TYPE "UDT_SDC_EMS_TS_COM"
VERSION : 0.1
   STRUCT
      VAL : "UDT_SDC_TS_IF_COMMAND_VAL";
      BIT : "UDT_SDC_TS_IF_COMMAND_BIT";
      FKT_SET : "UDT_SDC_EMS_FKT_BITs";
      FKT_RESET : "UDT_SDC_EMS_FKT_BITs";
   END_STRUCT;
END_TYPE

TYPE "UDT_EMS_IF_Q_STAT"
VERSION : 0.1
   STRUCT
      LIFE_BIT : Bool;   // Lebensbit / Heartbeat
      ER_SUM : Bool;   // Sammelfehler / Summaryerror
      IR_MAN : Bool;   // EMS in Handbetrieb / EMS in manual mode (IR)
      ER_RESET : Bool;   // Störung quittieren / Error reset (IR)
      HOIST_CLEAR : Bool;   // Hub über/in Sollpos und Bereit ohne Störung / Hoist above position and no error
      POS_START_X : Bool;   // Fahrantrieb positioniert / Drive positioning started
      ALWAYS_ONE : Bool;   // immer "1" / Always "1"
      H_DISABLED : Bool;   // Hub gesperrt / Hoist disabled
      D_FWD : Bool;   // Fahrantrieb fährt vorwärts / Drive moves forwards
      D_RWD : Bool;   // Fahrantrieb fährt rückwärts / Drive moves reward
      bit12 : Bool;   // Reserve / spare
      D_IN_POS : Bool;   // Fahrantrieb in Position / Drive in Position
      H_UP : Bool;   // Hub hebt / Hoist raises
      H_DOWN : Bool;   // Hub senkt / Hoist lowers
      H_IN_POS : Bool;   // Hub in Position / Hoist in position
      H_IN_TOPPOS : Bool;   // Hub in oberster Position / Hoist in top position
      bit2_0 : Bool;   // Schwenkantrieb fährt + / Tilt moves clockwise
      bit2_1 : Bool;   // Schwenkantrieb fährt - / Tilt moves counterclockwise
      bit2_2 : Bool;   // Hub in oberster Position / Tilt in position
      bit2_3 : Bool;   // Hub in Grundstellung / Tilt in home position
      IN_BOTPOS : Bool;   // Hub in unterster Position / Hoist In bottom Position (min) (with Tiltposition)
      bit2_5 : Bool;   // Reserve / spare
      bit2_6 : Bool;   // Reserve / spare
      bit2_7 : Bool;   // Reserve / spare
      MESS_ACT : Bool;   // Störnummer ist eine Meldung / Error No is a Message
      MESS_POS : Bool;   // Reserve / spare
      bit3_2 : Bool;   // Reserve / spare
      bit3_3 : Bool;   // Reserve / spare
      bit3_4 : Bool;   // Reserve / spare
      bit3_5 : Bool;   // Reserve / spare
      bit3_6 : Bool;   // Reserve / spare
      DATA_TRANS : Bool;   // Datentransfer ist aktiv / Data Transfer aktiv
   END_STRUCT;
END_TYPE

TYPE "UDT_EMS_IF_I_CONTR"
VERSION : 0.1
   STRUCT
      LIFE_BIT : Bool;   // Lebensbit / Heartbeat
      ER_SDC : Bool;   // Sammelfehler / Summaryerror
      H_EMERG : Bool;   // Hubantrieb Notbetrieb / Hoist Emergency mode
      Spare_0_3 : Bool;   // Schwenkantrieb Notbetrieb / Tilt Emergency mode
      LAMP_TEST : Bool;   // Lampentest / Lamp Test
      VAC_CLEAN : Bool;   // EMS mit Staubsauger / EMS with vac cleaner
      SYNCH : Bool;   // Synchronbetrieb / Control distance, synchronous area
      DATA_TRANS : Bool;   // Datentransfer ist aktiv / Data Transfer aktiv
      ER_RESET : Bool;   // Störung quittieren / Error reset
      AUTO : Bool;   // 1 = Automatikbetrieb / Automatic mode in section
      MAN : Bool;   // 1 = Handbetrieb / Manual mode in section
      D_C_BREAK : Bool;   // Fahrantrieb Befehl Bremse lüften / DRIVE Command release Break
      H_C_BREAK : Bool;   // Hubantrieb Befehl Bremse lüften / HOIST Command release Break
      D_EMERG_FC : Bool;   // Fahrantrieb Notbetrieb 1 Motor / DRIVE Emergency mode Frequencyconverter 1 Motor
      INC_TOL_POS : Bool;   // Schwenkantrieb Notbetrieb 1 Motor / TILT Emergency mode Frequencyconverter 1 Motor
      E_STOP : Bool;   // "1"Not-Halt / Emergency stop from Interface
      D_C_FWD : Bool;   // Fahrantrieb Befehl vorwärts / DRIVE Command forward
      D_C_RWD : Bool;   // Fahrantrieb Befehl rückwärts / DRIVE Command reward
      D_C_BSP : Bool;   // Fahrantrieb Befehl weiter fahren / DRIVE Command bridge stop position
      Spare_2_3 : Bool;   // Reserve / spare
      IR_noEMSnumber : Bool;   // Schwenkantrieb Befehl + / TILT Command clockwise
      IR_noLogin : Bool;   // Schwenkantrieb Befehl - / TILT Command counterclockwise
      BYP_scalance_PN_error : Bool;   // Schwenkantrieb Befehl positionieren / TILT Command positioning
      Spare_2_7 : Bool;   // Schwenkantrieb Befehl fahren in Grundstellung / TILT Command to home position, high priority
      H_C_UP : Bool;   // Hubantrieb Befehl heben / HOIST Command raise without positioning
      H_C_DOWN : Bool;   // Hubantrieb Befehl senken / HOIST Command lower without positioning
      H_C_POS : Bool;   // Hubantrieb Befehl positionieren / HOIST Command hoist positioning
      H_C_TOP : Bool;   // Hubantrieb Befehl fahren in oberste Position / HOIST Command Raise to top position, high priority
      H_EN : Bool;   // Hub-Schwenkfreigabe / HOIST-TILT enable
      H_BYP_ROPE : Bool;   // Überbrücken Seilkontrolle / Bypass monitoring of rope
      Spare_3_6 : Bool;   // Reserve / spare
      H_BYP_REF_INI : Bool;   // Überbrücken Kontrolle Referenzinitiator (nicht safety) / No monitoring of reference initiator (non safety)
   END_STRUCT;
END_TYPE

TYPE "UDT_SDC_TS_IF_COMMAND_BIT"
AUTHOR : SIEMENS
FAMILY : FT
NAME : SDC_BIT
VERSION : 2.0
   STRUCT
      ER_RESET : Bool;   // Error Reset
      AUTO : Bool;   // 1 = Automatik in Sektion
      MAN : Bool;   // 1 = Handbetrieb in Sektion
      Spare_0_3 : Bool;   // Reserve
      Spare_0_4 : Bool;   // Reserve
      E_STOP : Bool;   // "1" -> NotAus von Interface (system PLC)
      Spare_0_6 : Bool;   // Reserve
      Spare_0_7 : Bool;   // Reserve
      D_C_FWD : Bool;   // Fahrantrieb Kommando vorwärts
      D_C_RWD : Bool;   // Fahrantrieb Kommando rückwärts
      D_C_BSP : Bool;   // Fahrantrieb Kommando Überbrückung Stopp-Position
      D_C_V1 : Bool;   // Fahrantrieb Kommando Geschwindigkeit 1
      D_C_V2 : Bool;   // Fahrantrieb Kommando Geschwindigkeit 2
      D_C_V_VAR : Bool;   // Fahrantrieb Kommando variabler Geschwindigkeit
      D_C_BEFOR_POS : Bool;   // Fahrantrieb Kommando Freigabe vor Stop-Position
      D_C_AFTER_POS : Bool;   // Fahrantrieb Kommando Freigabe nach Stop-Position
      H_C_RAISE : Bool;   // Hubantrieb Kommando aufwärts
      H_C_LOWER : Bool;   // Hubantrieb Kommando abwärts
      H_C_POS : Bool;   // Hubantrieb Kommando Positionieren
      H_C_POS1 : Bool;   // Hubantrieb Kommando Offset 1
      H_C_POS2 : Bool;   // Hubantrieb Kommando Offset 2
      H_C_POS3 : Bool;   // Hubantrieb Kommando Offset 3
      H_C_POS4 : Bool;   // Hubantrieb Kommando Offset 4
      H_C_TOP : Bool;   // Hubantrieb Kommando nach Top Position, hohe Priorität
      H_BYP_ROPE : Bool;   // Hubantrieb Überbrücken Seilkontrolle
      Spare_3_1 : Bool;   // Reserve
      H_BYP_REF_INI : Bool;   // Hubantrieb Überbrücken Kontrolle Referenzinitiator (nicht safety)
      H_C_SLOW : Bool;   // Hubantrieb Kommando globaler Parameter langsam
      D_BYP_DIST_CONTR : Bool;   // Fahrantrieb Überbrücke Distanzkontrolle
      Spare_3_5 : Bool;   // Reserve
      Spare_3_6 : Bool;   // Reserve
      SET_PROF : Bool;   // setze Profile
   END_STRUCT;
END_TYPE

TYPE "UDT_SDC_TS_IF_COMMAND_VAL"
AUTHOR : SIEMENS
FAMILY : FT
NAME : SDC_VAL
VERSION : 1.6
   STRUCT
      PROFIL : Int;   // Profile
      D_SETSPEED : DInt;   // set value: drive speed (mm/min)
      D_POS_OFFS : Int;   // Antriebsposition offset
      H_POS_OFFS : Int;
   END_STRUCT;
END_TYPE

TYPE "UDT_SDC_TS_IF_STATUS_BIT"
AUTHOR : SIEMENS
FAMILY : FT
NAME : SDC_BIT
VERSION : 1.6
   STRUCT
      PRESENT : Bool;   // EMS vorhanden
      ERROR : Bool;   // Sammelstörung
      MAN_IR : Bool;   // EMS in Handbetrieb (Fernsteuerung)
      MORE_EMS_PRESENT : Bool;   // Mehr als 1 EMS in Sektion vorhanden
      ER_COMMAND : Bool;   // Fehlerhafte Befehle von System PLC
      W_DIST : Bool;   // Warnung Distanckontrolle ist aktiv
      Spare_0_6 : Bool;   // Warnung Auffahrsensor ist aktiv Reserve
      MESS_ACT : Bool;   // Störnummer ist eine Meldung / Error No is a Message
      D_MOVING : Bool;   // Fahrantrieb ist ein
      D_NOT_MOVING : Bool;   // Fahrantrieb ist aus
      H_MOVING : Bool;   // Hubantrieb ist ein
      H_NOT_MOVING : Bool;   // Hubantrieb ist aus
      X_MOVING : Bool;   // Reserve Antrieb ein
      X_NOT_MOVING : Bool;   // Reserve Antrieb aus
      D_IN_POS : Bool;   // Fahrantrieb in Position
      Spare_2_1 : Bool;   // Reserve
      D_BEFOR_POS : Bool;   // Fahrantrieb vor Stopposition
      D_AFTER_POS : Bool;   // Fahrantrieb nach Stopposition
      D_GR_AP1 : Bool;   // Fahrantrieb Barcodeposition größer Aktionspunkt 1
      D_SM_AP1 : Bool;   // Fahrantrieb Barcodeposition kleiner Aktionspunkt 1
      D_GR_AP2 : Bool;   // Fahrantrieb Barcodeposition größer Aktionspunkt 2
      D_SM_AP2 : Bool;   // Fahrantrieb Barcodeposition kleiner Aktionspunkt 2
      H_IN_POS : Bool;   // Hubantrieb in Position (hoist drive)
      H_IN_TOPPOS : Bool;   // Hubantrieb in top pos.(limit)
      H_IN_POS1 : Bool;   // Hubantrieb in Position (hoist drive) Offset 1
      H_IN_POS2 : Bool;   // Hubantrieb in Position (hoist drive) Offset 2
      H_IN_POS3 : Bool;   // Hubantrieb in Position (hoist drive) Offset 3
      H_IN_POS4 : Bool;   // Hubantrieb in Position (hoist drive) Offset 4
      H_GR_POS : Bool;   // Hubposition größer Sollposition ohne Offset
      H_SM_POS : Bool;   // Hubposition kleiner Sollposition ohne Offset
      H_GR_POS1 : Bool;   // Hubposition größer Sollposition + Offset 1
      H_SM_POS1 : Bool;   // Hubposition kleiner Sollposition + Offset 1
      H_GR_POS2 : Bool;   // Hubposition größer Sollposition + Offset 2
      H_SM_POS2 : Bool;   // Hubposition kleiner Sollposition + Offset 2
      H_GR_POS3 : Bool;   // Hubposition größer Sollposition + Offset 3
      H_SM_POS3 : Bool;   // Hubposition kleiner Sollposition + Offset 3
      H_GR_POS4 : Bool;   // Hubposition größer Sollposition + Offset 4
      H_SM_POS4 : Bool;   // Hubposition kleiner Sollposition + Offset 4
      H_BOTTOM_POS : Bool;   // Hub (mit Neigung) in unterer Position
      H_DISABLED : Bool;   // Hub ist verriegelt, keine Freigabe
      H_CLEAR : Bool;   // Hub über/in Sollpos und bereit ohne Störung
      D_MOVING_FWD : Bool;   // Fahrantrieb Bewegung vorwärts
      D_MOVING_RWD : Bool;   // Fahrantrieb Bewegung rückwärts
      D_RESET_AFTER : Bool;   // Fahrantrieb Bewegung Belegt Reset ohne Present
      D_PULK : Bool;   // Fahrantrieb Sektion in PULKbetrieb
      D_NO_POS : Bool;   // Fahrantrieb keine Stopposition Sektion
      Spare_7_6 : Bool;
      Spare_7_7 : Bool;
   END_STRUCT;
END_TYPE

TYPE "UDT_SDC_TS_IF_STATUS_VAL"
AUTHOR : SIEMENS
FAMILY : FT
NAME : SDC_VAL
VERSION : 1.6
   STRUCT
      EMS_ID : Int;   // EMS ID Nummer
      PROFIL : Int;   // Profile
      DRIVE_POS : DInt;   // Antriebsposition in mm
      HOIST_POS : Int;   // Höhe in mm
      ERROR : Int;   // Error-Nummer
      DRIVE_POS_PERC : Int;   // Position [% of Start End Section]
      SEK : Int;   // Sektion
   END_STRUCT;
END_TYPE

TYPE "UDT_SDC_EMS_FKT_BITs"
VERSION : 0.1
   STRUCT
      EMS_TO_REPAIR_1 : Bool;   // EMS zur Reperatur 1
      EMS_TO_REPAIR_2 : Bool;   // EMS zur Reperatur 2
      EMERG_HOIST : Bool;   // EMS Emergancy without Hoist
      Reserve_03 : Bool;   // EMS Emergancy without Tilt
      EMERG_DRIVE_FC : Bool;   // EMS Drive Emergency mode Frequencyconverter 1 Motor
      Reserve_05 : Bool;   // EMS Tilt Emergency mode Frequencyconverter 1 Motor
      LAMP_TEST : Bool;   // EMS Lamp Test
      VAC_CLEAN : Bool;   // EMS VAC Reiniger
      PE_TEST : Bool;   // EMS PE Test NIO
      KOHLE_TEST : Bool;   // EMS KOHLE Test NIO
      KOM_TEST : Bool;   // Reserve
      Reserve_11 : Bool;   // Reserve
      Reserve_12 : Bool;   // Reserve
      Reserve_13 : Bool;   // Reserve
      Reserve_14 : Bool;   // Reserve
      Reserve_15 : Bool;   // Reserve
   END_STRUCT;
END_TYPE

TYPE "UDT_EMS_IF_I_SDC_ERRORS"
VERSION : 0.1
   STRUCT
      _901_ER_SUM : Bool;   // Error SDC + EMS Summary
      _902_ER_SUM_SDC : Bool;   // Error SDC Summary
      _903_ER_BC_JUMP : Bool;   // Error SDC Barcode Jump
      _904_ER_NO_SEK : Bool;   // Error SDC no Section found
      _905_ER_COMMAND : Bool;   // Error SDC worng Commands from Main Plc
      _906_ER_BC_LIM : Bool;   // Error SDC Barcode LIMIT
      _907_ER_EMS_ID : Bool;   // Error SDC wrong EMS Number
      _908_ER_SEK_NR : Bool;   // Error SDC wrong Sektion Number
      _909_ER_LIFE : Bool;   // Error SDC Lifebeat to EMS
      _910_ER_BUS : Bool;   // Error SDC no Buscommunication to EMS device
      _911 : Bool;   // spare
      _912 : Bool;   // spare
      _913 : Bool;   // spare
      _914 : Bool;   // spare
      _915 : Bool;   // spare
      _916 : Bool;   // spare
   END_STRUCT;
END_TYPE

TYPE "UDT_SDC_ERROR_STAT"
VERSION : 0.1
   STRUCT
      EMS_TS_STAT_VAL : "UDT_SDC_TS_IF_STATUS_VAL";
      ER : "UDT_EMS_IF_I_SDC_ERRORS";
      Spare : Int;   // spare
      ER_DATE : Date_And_Time;   // Fehler Zeit
   END_STRUCT;
END_TYPE

// folder: UDT_AB_Interlocks

TYPE "UDT_AB_Interlocks_Carrier"
VERSION : 0.1
   STRUCT
      Carrier_IN : "UDT_AB_Interlocks_Carrier_In";
      Carrier_OUT : "UDT_AB_Interlocks_Carrier_Out";
   END_STRUCT;
END_TYPE

TYPE "UDT_AB_Interlocks_SDC_In"
VERSION : 0.1
   STRUCT
      EMS01_MasterPowerOn : Bool;
      EMS01_Fault_Reset_PB : Bool;
      EMS01R1_MasterPowerOn : Bool;
      EMS01R1_Fault_Reset_PB : Bool;
      EMS01R2_MasterPowerOn : Bool;
      EMS01R2_Fault_Reset_PB : Bool;
      EMS01R3_MasterPowerOn : Bool;
      EMS01R3_Fault_Reset_PB : Bool;
      EMS01R4_MasterPowerOn : Bool;
      EMS01R4_Fault_Reset_PB : Bool;
      EMS_Stop_26_Set_To_Release : Bool;
      Spare_11 : Bool;
      Spare_12 : Bool;
      Spare_13 : Bool;
      Spare_14 : Bool;
      Heartbeat : Bool;
      SpareWord2 : Word;
      SpareWord3 : Word;
      CarrierSpeedRef : Word;
      ProductionSpeedRef : Word;
   END_STRUCT;
END_TYPE

TYPE "UDT_AB_Interlocks_CarrierStatus_Out"
VERSION : 0.1
   STRUCT
      Spare0 : Bool;
      DriveTripped : Bool;
      Spare2 : Bool;
      PositioningComplete : Bool;
      RunStopPressed : Bool;
      Moving : Bool;
      Faulted : Bool;
      InAuto : Bool;
      Spare8 : Bool;
      Spare9 : Bool;
      Spare10 : Bool;
      Spare11 : Bool;
      Spare12 : Bool;
      Spare13 : Bool;
      Spare14 : Bool;
      Spare15 : Bool;
   END_STRUCT;
END_TYPE

TYPE "UDT_AB_Interlocks_Carrier_Out"
VERSION : 0.1
   STRUCT
      Status : "UDT_AB_Interlocks_CarrierStatus_Out";
      Fault : Word;
      Position : DWord;
      Zone : Word;
   END_STRUCT;
END_TYPE

TYPE "UDT_AB_Interlocks_Carrier_In"
VERSION : 0.1
   STRUCT
      CarrierDelete : Bool;
   END_STRUCT;
END_TYPE

TYPE "UDT_AB_Interlocks"
VERSION : 0.1
   STRUCT
      SDC_Interlocks_In : "UDT_AB_Interlocks_SDC_In";
      SDC_Interlocks_Out : "UDT_AB_Interlocks_SDC_Out";
      Carrier : Array[1..99] of "UDT_AB_Interlocks_Carrier";
   END_STRUCT;
END_TYPE

TYPE "UDT_AB_Interlocks_SDC_Out"
VERSION : 0.1
   STRUCT
      SDC_Faulted : Bool;
      SDC_Status_1 : Bool;
      SDC_Status_2 : Bool;
      SDC_Status_3 : Bool;
      SDC_Status_4 : Bool;
      SDC_Status_5 : Bool;
      SDC_Status_6 : Bool;
      SDC_Status_7 : Bool;
      SDC_Status_8 : Bool;
      SDC_Status_9 : Bool;
      SDC_Status_10 : Bool;
      SDC_Status_11 : Bool;
      SDC_Status_12 : Bool;
      SDC_Status_13 : Bool;
      SDC_Status_14 : Bool;
      Heartbeat : Bool;
   END_STRUCT;
END_TYPE

// folder: UserDiag

TYPE "UserDiag_typeDevice"
TITLE = UserDiag_typeDevice
VERSION : 0.1
   STRUCT
      hardwareId : Hw_Device := 16#0000;   // Hardware identifier of the device/slave
      number : UInt := 0;   // Profinet device number/Profibus address of the slave
      "name" : String[50];   // Name of the device/slave
      ipAddress : IP_V4;   // IP address of the device
      state : USInt := 0;   // Status of the device/slave. 1:ok; 2:faulty, 3:lost connection, 4:disabled, 5:problem, 12:was faulty, 13:was lost, 14:was disabled, 15:problem gone
      exists : Bool := FALSE;   // TRUE: Device/slave is existing
      configured : Bool := FALSE;   // TRUE: Device/slave is configured
      faulty : Bool := FALSE;   // TRUE: Device/slave is faulty
      problem : Bool := FALSE;   // TRUE: Device/slave has a problem
      disabled : Bool := FALSE;   // TRUE: Device/slave is disabled
      error : Bool := FALSE;   // TRUE: Error in device/slave
      nextDevice : Int;   // device number of next device
      actualConfiguredSlots : Int := 0;   // Number of configured slots in the device/slave
      slots : Array[0.."USERDIAG_SLOTS_PER_DEVICE_UPPER_LIM"] of "UserDiag_typeSlot";   // Slot information of a device/slave
   END_STRUCT;
END_TYPE

TYPE "UserDiag_typeIOSystem"
TITLE = UserDiag_typeIOSystem
VERSION : 0.1
   STRUCT
      hardwareId : Hw_IoSystem := 16#0000;   // Hardware identifier of the IO-System/DP-Mastersystem
      number : UInt := 0;   // IO-System/DP-Mastersystem number
      error : Bool := FALSE;   // TRUE: Error in IO-System/DP-Mastersystem
      firstDevice : Int := 0;   // device number (index) of first device in IO System
      lastDevice : Int := 0;   // device number (index) of last device IO System
      actualConfiguredDevices : Int := 0;   // Number of configured devices/slaves in IO-System/DP-Mastersystem
      devices : Array[1.."USERDIAG_DEVICES_PER_IO_SYSTEM_UPPER_LIM"] of "UserDiag_typeDevice";   // Device/Slave information
   END_STRUCT;
END_TYPE

TYPE "UserDiag_typeActIOSystem"
TITLE = UserDiag_typeActIOSystem
VERSION : 0.1
   STRUCT
      actIOSystemNumber : Int := 1;   // Number of actual selected IO-system/DP-Mastersystem
      actIODeviceNumbers : Array[1.."USERDIAG_DEVICES_PER_SCREEN_UPPER_LIM"] of UInt;   // Device numbers/profibus addresses of actual selected IO-System/DP-Mastersystem
      actIODeviceState : Array[1.."USERDIAG_DEVICES_PER_SCREEN_UPPER_LIM"] of USInt;   // State of devices/slaves in actual selected IO-System/DP-Mastersystem
      actDeviceSlotsUsed : Array[0.."USERDIAG_SLOTS_PER_SCREEN_UPPER_LIM"] of Bool;   // Used slots of actual selected device/slave
      actDeviceSlotsState : Array[0.."USERDIAG_SLOTS_PER_SCREEN_UPPER_LIM"] of USInt;   // States of actual selected device/slave
   END_STRUCT;
END_TYPE

TYPE "UserDiag_typeHmiData"
VERSION : 0.1
   STRUCT
      actIOSystem : Int := 1;   // Index of actual selected IO-System/DP-Mastersystem
      actDeviceOfScreen : Int := 1;   // Index of selected device/slave on actual Screen
      ioSlotDiagnosticsLoaded : Bool;   // TRUE: Page for slot diagnostics is loaded
      actScreenDevices : Int := 1;   // Actual screennumber for copying device status to HMI
      maxScreensDevices : Int;   // Maximum screennumber for copying device status to HMI
      ackWaitTime : Int;   // Wait time after startup, for auto acknowledge
      ackStates : Bool;   // TRUE: Acknowledge of occurred errors in device/slave
      actIOSystemData : "UserDiag_typeActIOSystem";   // Data of actual IO system
      actDeviceNumber : UInt;   // Actual number/profibus address of device/slave
      actDeviceName : String[50];   // Name of actual selected device/slave
      actIPAddress : IP_V4;   // IP address of the device
      errorAtLowerScreen : Bool;   // Error at lower screen
      errorAtUpperScreen : Bool;   // Error at upper screen
      filterErrorDevices : Bool;   // Filter only fault devices
      ioSystemError : Array[1.."USERDIAG_IO_SYSTEMS_UPPER_LIM"] of Bool;   // Error in IO systems
   END_STRUCT;
END_TYPE

TYPE "UserDiag_typeSlot"
TITLE = UserDiag_typeSlot
VERSION : 0.1
   STRUCT
      hardwareId : Hw_Io := 16#0000;   // Hardware identifier of the module which is inserted in the slot
      state : USInt := 0;   // Status of the device/slave. 1:ok; 2:faulty, 3:lost connection, 4:disabled, 5:problem, 12:was faulty, 13:was lost, 14:was disabled, 15:problem gone
      exists : Bool := FALSE;   // TRUE: Modul is existing
      configured : Bool := FALSE;   // TRUE: Modul is configured
      faulty : Bool := FALSE;   // TRUE: Modul is faulty
      problem : Bool := FALSE;   // TRUE: Modul has a problem
      disabled : Bool := FALSE;   // TRUE: Modul is disabled
      error : Bool := FALSE;   // TRUE: Error in module which is inserted in the slot
   END_STRUCT;
END_TYPE

TYPE "UserDiag_typePLC"
TITLE = UserDiag_typePLC
VERSION : 0.1
   STRUCT
      hardwareId : Hw_Device := 16#0000;   // Hardware identifier of the PLC
      error : Bool := FALSE;   // TRUE: Error in PLC
      actualConfiguredSlots : Int := 0;   // Number of configured local slots at PLC
      slots : Array[0.."USERDIAG_SLOTS_PER_PLC_UPPER_LIM"] of "UserDiag_typeSlot";   // Information of the PLC slots; index = slotnumber; PLC always at slot 1
   END_STRUCT;
END_TYPE

// folder: 04_FCs

DATA_BLOCK "IDB558_ZONE_07"   // DB13
{ S7_Optimized_Access := 'FALSE' }
VERSION : 0.1
"FB115_FB_Zone"
BEGIN
END_DATA_BLOCK

// folder: 05_DBs

DATA_BLOCK "DB_SDC_TS_IF_COM_LOE"   // DB4
{ S7_Optimized_Access := 'FALSE' }
VERSION : 0.1
   VAR
      LoeSEK : "UDT_SDC_EMS_TS_COM";
   END_VAR
BEGIN
END_DATA_BLOCK

DATA_BLOCK "EMS"   // DB8
{ S7_Optimized_Access := 'TRUE' }
VERSION : 0.1
BEGIN
   Production_Spacing := 1000;
   Carrier_Spacing := 800;
END_DATA_BLOCK

DATA_BLOCK "DB11_CARRIER"   // DB11
{ S7_Optimized_Access := 'TRUE' }
VERSION : 0.1
BEGIN
END_DATA_BLOCK

DATA_BLOCK "DB14_CarrZnFindArrayBuffer"   // DB14
{ S7_Optimized_Access := 'TRUE' }
VERSION : 0.1
BEGIN
END_DATA_BLOCK

DATA_BLOCK "DB15__FB_Zone_DB"   // DB15
{ S7_Optimized_Access := 'FALSE' }
VERSION : 0.1
"FB115_FB_Zone"
BEGIN
END_DATA_BLOCK

DATA_BLOCK "DB16_EMS_Status"   // DB16
{ S7_Optimized_Access := 'TRUE' }
VERSION : 0.1
   VAR
      EMS_DeviceStates : Struct
         Profinet1_Lddr : Hw_IoSystem := 257;
         DeviceStates_Mode2 : UInt := 2;
         DeviceStates_Mode4 : UInt := 4;
         DeviceStates_Mode5 : UInt := 5;
         DeviceStates_RetVal_2 : Int;
         DeviceStates_RetVal_4 : Int;
         DeviceStates_RetVal_5 : Int;
         DeviceStates_State2 : Array[0..1023] of Bool;
         DeviceStates_State4 : Array[0..1023] of Bool;
         DeviceStates_State5 : Array[0..1023] of Bool;
         DeviceStates_Condition_HMI : Array[0..82] of Int;
      END_STRUCT;
   END_VAR
BEGIN
END_DATA_BLOCK

DATA_BLOCK "TC_SDC_Out"   // DB53
{ S7_Optimized_Access := 'TRUE' }
VERSION : 0.1
BEGIN
END_DATA_BLOCK

DATA_BLOCK "DB101_DB_SDC_FAULTS"   // DB101
{ S7_Optimized_Access := 'FALSE' }
VERSION : 0.1
   VAR
      SDC_Fault : Word;
      Carrier_Fault : Array[1..90] of Word;
   END_VAR
BEGIN
END_DATA_BLOCK

DATA_BLOCK "DB110_DB_SDC_IN"   // DB110
{ S7_Optimized_Access := 'TRUE' }
VERSION : 0.1
   VAR
      Carrier : Array[0..99] of "UDT_SDC_IN";
   END_VAR
BEGIN
END_DATA_BLOCK

DATA_BLOCK "DB111_DB_SDC_OUT"   // DB111
{ S7_Optimized_Access := 'TRUE' }
VERSION : 0.1
   VAR
      Carrier : Array[0..99] of "UDT_SDC_OUT";
   END_VAR
BEGIN
END_DATA_BLOCK

DATA_BLOCK "DB116_TC_ZoneMotionControl"   // DB116
{ S7_Optimized_Access := 'TRUE' }
VERSION : 0.1
BEGIN
END_DATA_BLOCK

DATA_BLOCK "DB302_HMI_Faults"   // DB302
{ S7_Optimized_Access := 'TRUE' }
VERSION : 0.1
   VAR
      SDC_Faults_0 : Int := 0;
      SDC_Faults_1 : Int := 0;
      SDC_Faults_2 : Int := 0;
      SDC_Faults_3 : Int := 0;
      Carrier1_Faults_0 : Int := 0;
      Carrier1_Faults_1 : Int := 0;
      Carrier1_Faults_2 : Int := 0;
      Carrier1_Faults_3 : Int := 0;
      Carrier2_Faults_0 : Int := 0;
      Carrier2_Faults_1 : Int := 0;
      Carrier2_Faults_2 : Int := 0;
      Carrier2_Faults_3 : Int := 0;
      Carrier3_Faults_0 : Int := 0;
      Carrier3_Faults_1 : Int := 0;
      Carrier3_Faults_2 : Int := 0;
      Carrier3_Faults_3 : Int := 0;
      Carrier4_Faults_0 : Int := 0;
      Carrier4_Faults_1 : Int := 0;
      Carrier4_Faults_2 : Int := 0;
      Carrier4_Faults_3 : Int := 0;
      Carrier5_Faults_0 : Int := 1;
      Carrier5_Faults_1 : Int := 2;
      Carrier5_Faults_2 : Int := 3;
      Carrier5_Faults_3 : Int := 4;
      Carrier6_Faults_0 : Int := 5;
      Carrier6_Faults_1 : Int := 6;
      Carrier6_Faults_2 : Int := 7;
      Carrier6_Faults_3 : Int := 8;
      Carrier7_Faults_0 : Int := 9;
      Carrier7_Faults_1 : Int := 10;
      Carrier7_Faults_2 : Int := 11;
      Carrier7_Faults_3 : Int := 12;
      Carrier8_Faults_0 : Int := 13;
      Carrier8_Faults_1 : Int := 14;
      Carrier8_Faults_2 : Int := 15;
      Carrier8_Faults_3 : Int := 16;
      Carrier9_Faults_0 : Int := 17;
      Carrier9_Faults_1 : Int := 18;
      Carrier9_Faults_2 : Int := 19;
      Carrier9_Faults_3 : Int := 20;
      Carrier10_Faults_0 : Int := 21;
      Carrier10_Faults_1 : Int := 22;
      Carrier10_Faults_2 : Int := 23;
      Carrier10_Faults_3 : Int := 24;
      Carrier11_Faults_0 : Int := 25;
      Carrier11_Faults_1 : Int := 26;
      Carrier11_Faults_2 : Int := 27;
      Carrier11_Faults_3 : Int := 28;
      Carrier12_Faults_0 : Int := 29;
      Carrier12_Faults_1 : Int := 30;
      Carrier12_Faults_2 : Int := 31;
      Carrier12_Faults_3 : Int := 32;
      Carrier13_Faults_0 : Int := 33;
      Carrier13_Faults_1 : Int := 34;
      Carrier13_Faults_2 : Int := 35;
      Carrier13_Faults_3 : Int := 36;
      Carrier14_Faults_0 : Int := 37;
      Carrier14_Faults_1 : Int := 38;
      Carrier14_Faults_2 : Int := 39;
      Carrier14_Faults_3 : Int := 40;
      Carrier15_Faults_0 : Int := 41;
      Carrier15_Faults_1 : Int := 42;
      Carrier15_Faults_2 : Int := 43;
      Carrier15_Faults_3 : Int := 44;
      Carrier16_Faults_0 : Int := 45;
      Carrier16_Faults_1 : Int := 46;
      Carrier16_Faults_2 : Int := 47;
      Carrier16_Faults_3 : Int := 48;
      Carrier17_Faults_0 : Int := 49;
      Carrier17_Faults_1 : Int := 50;
      Carrier17_Faults_2 : Int := 51;
      Carrier17_Faults_3 : Int := 52;
      Carrier18_Faults_0 : Int := 53;
      Carrier18_Faults_1 : Int := 54;
      Carrier18_Faults_2 : Int := 55;
      Carrier18_Faults_3 : Int := 56;
      Carrier19_Faults_0 : Int := 57;
      Carrier19_Faults_1 : Int := 58;
      Carrier19_Faults_2 : Int := 59;
      Carrier19_Faults_3 : Int := 60;
      Carrier20_Faults_0 : Int := 61;
      Carrier20_Faults_1 : Int := 62;
      Carrier20_Faults_2 : Int := 63;
      Carrier20_Faults_3 : Int := 64;
      Carrier21_Faults_0 : Int := 65;
      Carrier21_Faults_1 : Int := 66;
      Carrier21_Faults_2 : Int := 67;
      Carrier21_Faults_3 : Int := 68;
      Carrier22_Faults_0 : Int := 69;
      Carrier22_Faults_1 : Int := 70;
      Carrier22_Faults_2 : Int := 71;
      Carrier22_Faults_3 : Int := 72;
      Carrier23_Faults_0 : Int := 73;
      Carrier23_Faults_1 : Int := 74;
      Carrier23_Faults_2 : Int := 75;
      Carrier23_Faults_3 : Int := 76;
      Carrier24_Faults_0 : Int := 77;
      Carrier24_Faults_1 : Int := 78;
      Carrier24_Faults_2 : Int := 79;
      Carrier24_Faults_3 : Int := 80;
      Carrier25_Faults_0 : Int := 81;
      Carrier25_Faults_1 : Int := 82;
      Carrier25_Faults_2 : Int := 83;
      Carrier25_Faults_3 : Int := 84;
      Carrier26_Faults_0 : Int := 85;
      Carrier26_Faults_1 : Int := 86;
      Carrier26_Faults_2 : Int := 87;
      Carrier26_Faults_3 : Int := 88;
      Carrier27_Faults_0 : Int := 89;
      Carrier27_Faults_1 : Int := 90;
      Carrier27_Faults_2 : Int := 91;
      Carrier27_Faults_3 : Int := 92;
      Carrier28_Faults_0 : Int := 93;
      Carrier28_Faults_1 : Int := 94;
      Carrier28_Faults_2 : Int := 95;
      Carrier28_Faults_3 : Int := 96;
      Carrier29_Faults_0 : Int := 97;
      Carrier29_Faults_1 : Int := 98;
      Carrier29_Faults_2 : Int := 99;
      Carrier29_Faults_3 : Int := 100;
      Carrier30_Faults_0 : Int := 101;
      Carrier30_Faults_1 : Int := 102;
      Carrier30_Faults_2 : Int := 103;
      Carrier30_Faults_3 : Int := 104;
      Carrier31_Faults_0 : Int := 105;
      Carrier31_Faults_1 : Int := 106;
      Carrier31_Faults_2 : Int := 107;
      Carrier31_Faults_3 : Int := 108;
      Carrier32_Faults_0 : Int := 109;
      Carrier32_Faults_1 : Int := 110;
      Carrier32_Faults_2 : Int := 111;
      Carrier32_Faults_3 : Int := 112;
      Carrier33_Faults_0 : Int := 113;
      Carrier33_Faults_1 : Int := 114;
      Carrier33_Faults_2 : Int := 115;
      Carrier33_Faults_3 : Int := 116;
      Carrier34_Faults_0 : Int := 117;
      Carrier34_Faults_1 : Int := 118;
      Carrier34_Faults_2 : Int := 119;
      Carrier34_Faults_3 : Int := 120;
      Carrier35_Faults_0 : Int := 121;
      Carrier35_Faults_1 : Int := 122;
      Carrier35_Faults_2 : Int := 123;
      Carrier35_Faults_3 : Int := 124;
      Carrier36_Faults_0 : Int := 125;
      Carrier36_Faults_1 : Int := 126;
      Carrier36_Faults_2 : Int := 127;
      Carrier36_Faults_3 : Int := 128;
      Carrier37_Faults_0 : Int := 129;
      Carrier37_Faults_1 : Int := 130;
      Carrier37_Faults_2 : Int := 131;
      Carrier37_Faults_3 : Int := 132;
      Carrier38_Faults_0 : Int := 133;
      Carrier38_Faults_1 : Int := 134;
      Carrier38_Faults_2 : Int := 135;
      Carrier38_Faults_3 : Int := 136;
      Carrier39_Faults_0 : Int := 137;
      Carrier39_Faults_1 : Int := 138;
      Carrier39_Faults_2 : Int := 139;
      Carrier39_Faults_3 : Int := 140;
      Carrier40_Faults_0 : Int := 141;
      Carrier40_Faults_1 : Int := 142;
      Carrier40_Faults_2 : Int := 143;
      Carrier40_Faults_3 : Int := 144;
      Carrier41_Faults_0 : Int := 145;
      Carrier41_Faults_1 : Int := 146;
      Carrier41_Faults_2 : Int := 147;
      Carrier41_Faults_3 : Int := 148;
      Carrier42_Faults_0 : Int := 149;
      Carrier42_Faults_1 : Int := 150;
      Carrier42_Faults_2 : Int := 151;
      Carrier42_Faults_3 : Int := 152;
      Carrier43_Faults_0 : Int := 153;
      Carrier43_Faults_1 : Int := 154;
      Carrier43_Faults_2 : Int := 155;
      Carrier43_Faults_3 : Int := 156;
      Carrier44_Faults_0 : Int := 157;
      Carrier44_Faults_1 : Int := 158;
      Carrier44_Faults_2 : Int := 159;
      Carrier44_Faults_3 : Int := 160;
      Carrier45_Faults_0 : Int := 161;
      Carrier45_Faults_1 : Int := 162;
      Carrier45_Faults_2 : Int := 163;
      Carrier45_Faults_3 : Int := 164;
      Carrier46_Faults_0 : Int := 165;
      Carrier46_Faults_1 : Int := 166;
      Carrier46_Faults_2 : Int := 167;
      Carrier46_Faults_3 : Int := 168;
      Carrier47_Faults_0 : Int := 169;
      Carrier47_Faults_1 : Int := 170;
      Carrier47_Faults_2 : Int := 171;
      Carrier47_Faults_3 : Int := 172;
      Carrier48_Faults_0 : Int := 173;
      Carrier48_Faults_1 : Int := 174;
      Carrier48_Faults_2 : Int := 175;
      Carrier48_Faults_3 : Int := 176;
      Carrier49_Faults_0 : Int := 177;
      Carrier49_Faults_1 : Int := 178;
      Carrier49_Faults_2 : Int := 179;
      Carrier49_Faults_3 : Int := 180;
      Carrier50_Faults_0 : Int := 181;
      Carrier50_Faults_1 : Int := 182;
      Carrier50_Faults_2 : Int := 183;
      Carrier50_Faults_3 : Int := 184;
      Carrier51_Faults_0 : Int := 185;
      Carrier51_Faults_1 : Int := 186;
      Carrier51_Faults_2 : Int := 187;
      Carrier51_Faults_3 : Int := 188;
      Carrier52_Faults_0 : Int := 189;
      Carrier52_Faults_1 : Int := 190;
      Carrier52_Faults_2 : Int := 191;
      Carrier52_Faults_3 : Int := 192;
      Carrier53_Faults_0 : Int := 193;
      Carrier53_Faults_1 : Int := 194;
      Carrier53_Faults_2 : Int := 195;
      Carrier53_Faults_3 : Int := 196;
      Carrier54_Faults_0 : Int := 197;
      Carrier54_Faults_1 : Int := 198;
      Carrier54_Faults_2 : Int := 199;
      Carrier54_Faults_3 : Int := 200;
      Carrier55_Faults_0 : Int := 201;
      Carrier55_Faults_1 : Int := 202;
      Carrier55_Faults_2 : Int := 203;
      Carrier55_Faults_3 : Int := 204;
      Carrier56_Faults_0 : Int := 205;
      Carrier56_Faults_1 : Int := 206;
      Carrier56_Faults_2 : Int := 207;
      Carrier56_Faults_3 : Int := 208;
      Carrier57_Faults_0 : Int := 209;
      Carrier57_Faults_1 : Int := 210;
      Carrier57_Faults_2 : Int := 211;
      Carrier57_Faults_3 : Int := 212;
      Carrier58_Faults_0 : Int := 213;
      Carrier58_Faults_1 : Int := 214;
      Carrier58_Faults_2 : Int := 215;
      Carrier58_Faults_3 : Int := 216;
      Carrier59_Faults_0 : Int := 217;
      Carrier59_Faults_1 : Int := 218;
      Carrier59_Faults_2 : Int := 219;
      Carrier59_Faults_3 : Int := 220;
      Carrier60_Faults_0 : Int := 221;
      Carrier60_Faults_1 : Int := 222;
      Carrier60_Faults_2 : Int := 223;
      Carrier60_Faults_3 : Int := 224;
      Carrier61_Faults_0 : Int := 225;
      Carrier61_Faults_1 : Int := 226;
      Carrier61_Faults_2 : Int := 227;
      Carrier61_Faults_3 : Int := 228;
      Carrier62_Faults_0 : Int := 229;
      Carrier62_Faults_1 : Int := 230;
      Carrier62_Faults_2 : Int := 231;
      Carrier62_Faults_3 : Int := 232;
      Carrier63_Faults_0 : Int := 233;
      Carrier63_Faults_1 : Int := 234;
      Carrier63_Faults_2 : Int := 235;
      Carrier63_Faults_3 : Int := 236;
      Carrier64_Faults_0 : Int := 237;